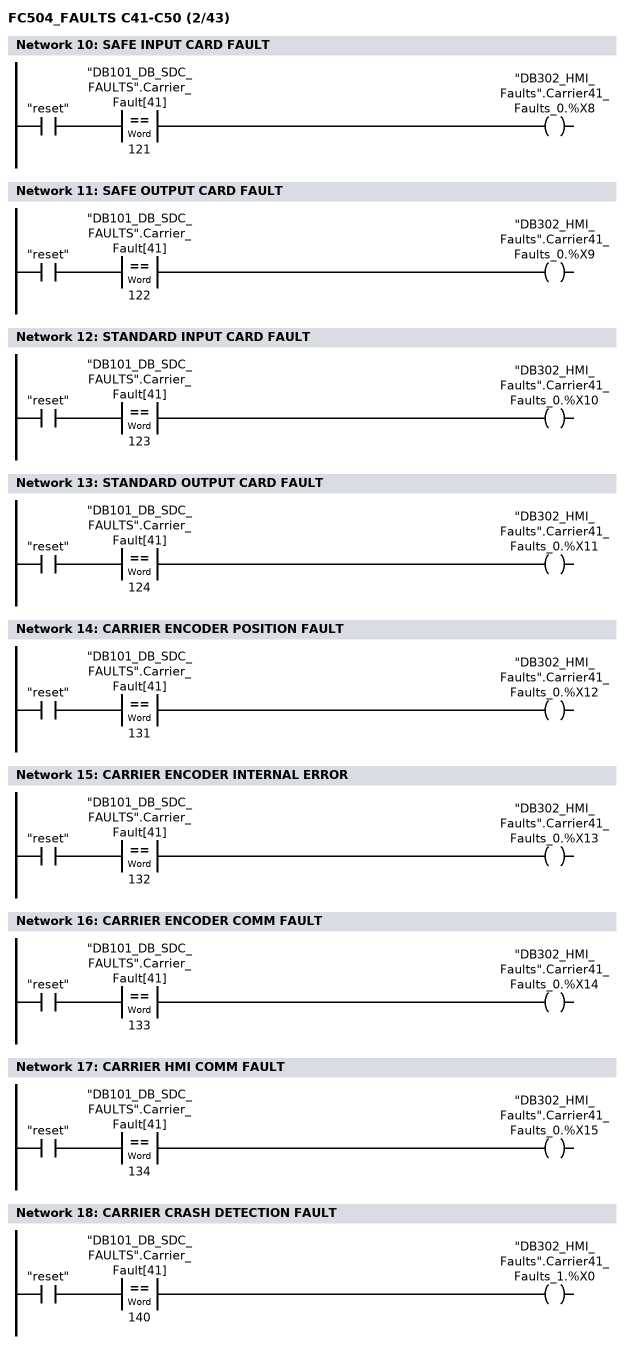
   RUNG wire#powerrail
      Contact( "reset" )
      { S7_Templates := "SrcType := Word" } EQ_Contact(in1 := "DB101_DB_SDC_FAULTS".Carrier_Fault[41], in2 := 121)
      Coil( "DB302_HMI_Faults".Carrier41_Faults_0.%X8 )
   END_RUNG
   // the same network as SCL:
   "DB302_HMI_Faults".Carrier41_Faults_0.%X8 := "reset" AND ("DB101_DB_SDC_FAULTS".Carrier_Fault[41] = 121);
END_REGION

REGION Network 11: SAFE OUTPUT CARD FAULT
   RUNG wire#powerrail
      Contact( "reset" )
      { S7_Templates := "SrcType := Word" } EQ_Contact(in1 := "DB101_DB_SDC_FAULTS".Carrier_Fault[41], in2 := 122)
      Coil( "DB302_HMI_Faults".Carrier41_Faults_0.%X9 )
   END_RUNG
   // the same network as SCL:
   "DB302_HMI_Faults".Carrier41_Faults_0.%X9 := "reset" AND ("DB101_DB_SDC_FAULTS".Carrier_Fault[41] = 122);
END_REGION

REGION Network 12: STANDARD INPUT CARD FAULT
   RUNG wire#powerrail
      Contact( "reset" )
      { S7_Templates := "SrcType := Word" } EQ_Contact(in1 := "DB101_DB_SDC_FAULTS".Carrier_Fault[41], in2 := 123)
      Coil( "DB302_HMI_Faults".Carrier41_Faults_0.%X10 )
   END_RUNG
   // the same network as SCL:
   "DB302_HMI_Faults".Carrier41_Faults_0.%X10 := "reset" AND ("DB101_DB_SDC_FAULTS".Carrier_Fault[41] = 123);
END_REGION

REGION Network 13: STANDARD OUTPUT CARD FAULT
   RUNG wire#powerrail
      Contact( "reset" )
      { S7_Templates := "SrcType := Word" } EQ_Contact(in1 := "DB101_DB_SDC_FAULTS".Carrier_Fault[41], in2 := 124)
      Coil( "DB302_HMI_Faults".Carrier41_Faults_0.%X11 )
   END_RUNG
   // the same network as SCL:
   "DB302_HMI_Faults".Carrier41_Faults_0.%X11 := "reset" AND ("DB101_DB_SDC_FAULTS".Carrier_Fault[41] = 124);
END_REGION

REGION Network 14: CARRIER ENCODER POSITION FAULT
   RUNG wire#powerrail
      Contact( "reset" )
      { S7_Templates := "SrcType := Word" } EQ_Contact(in1 := "DB101_DB_SDC_FAULTS".Carrier_Fault[41], in2 := 131)
      Coil( "DB302_HMI_Faults".Carrier41_Faults_0.%X12 )
   END_RUNG
   // the same network as SCL:
   "DB302_HMI_Faults".Carrier41_Faults_0.%X12 := "reset" AND ("DB101_DB_SDC_FAULTS".Carrier_Fault[41] = 131);
END_REGION

REGION Network 15: CARRIER ENCODER INTERNAL ERROR
   RUNG wire#powerrail
      Contact( "reset" )
      { S7_Templates := "SrcType := Word" } EQ_Contact(in1 := "DB101_DB_SDC_FAULTS".Carrier_Fault[41], in2 := 132)
      Coil( "DB302_HMI_Faults".Carrier41_Faults_0.%X13 )
   END_RUNG
   // the same network as SCL:
   "DB302_HMI_Faults".Carrier41_Faults_0.%X13 := "reset" AND ("DB101_DB_SDC_FAULTS".Carrier_Fault[41] = 132);
END_REGION

REGION Network 16: CARRIER ENCODER COMM FAULT
   RUNG wire#powerrail
      Contact( "reset" )
      { S7_Templates := "SrcType := Word" } EQ_Contact(in1 := "DB101_DB_SDC_FAULTS".Carrier_Fault[41], in2 := 133)
      Coil( "DB302_HMI_Faults".Carrier41_Faults_0.%X14 )
   END_RUNG
   // the same network as SCL:
   "DB302_HMI_Faults".Carrier41_Faults_0.%X14 := "reset" AND ("DB101_DB_SDC_FAULTS".Carrier_Fault[41] = 133);
END_REGION

REGION Network 17: CARRIER HMI COMM FAULT
   RUNG wire#powerrail
      Contact( "reset" )
      { S7_Templates := "SrcType := Word" } EQ_Contact(in1 := "DB101_DB_SDC_FAULTS".Carrier_Fault[41], in2 := 134)
      Coil( "DB302_HMI_Faults".Carrier41_Faults_0.%X15 )
   END_RUNG
   // the same network as SCL:
   "DB302_HMI_Faults".Carrier41_Faults_0.%X15 := "reset" AND ("DB101_DB_SDC_FAULTS".Carrier_Fault[41] = 134);
END_REGION

REGION Network 18: CARRIER CRASH DETECTION FAULT
   RUNG wire#powerrail
      Contact( "reset" )
      { S7_Templates := "SrcType := Word" } EQ_Contact(in1 := "DB101_DB_SDC_FAULTS".Carrier_Fault[41], in2 := 140)
      Coil( "DB302_HMI_Faults".Carrier41_Faults_1.%X0 )
   END_RUNG
   // the same network as SCL:
   "DB302_HMI_Faults".Carrier41_Faults_1.%X0 := "reset" AND ("DB101_DB_SDC_FAULTS".Carrier_Fault[41] = 140);
END_REGION

REGION Network 19: CARRIER NUMBER INVALID FAULT
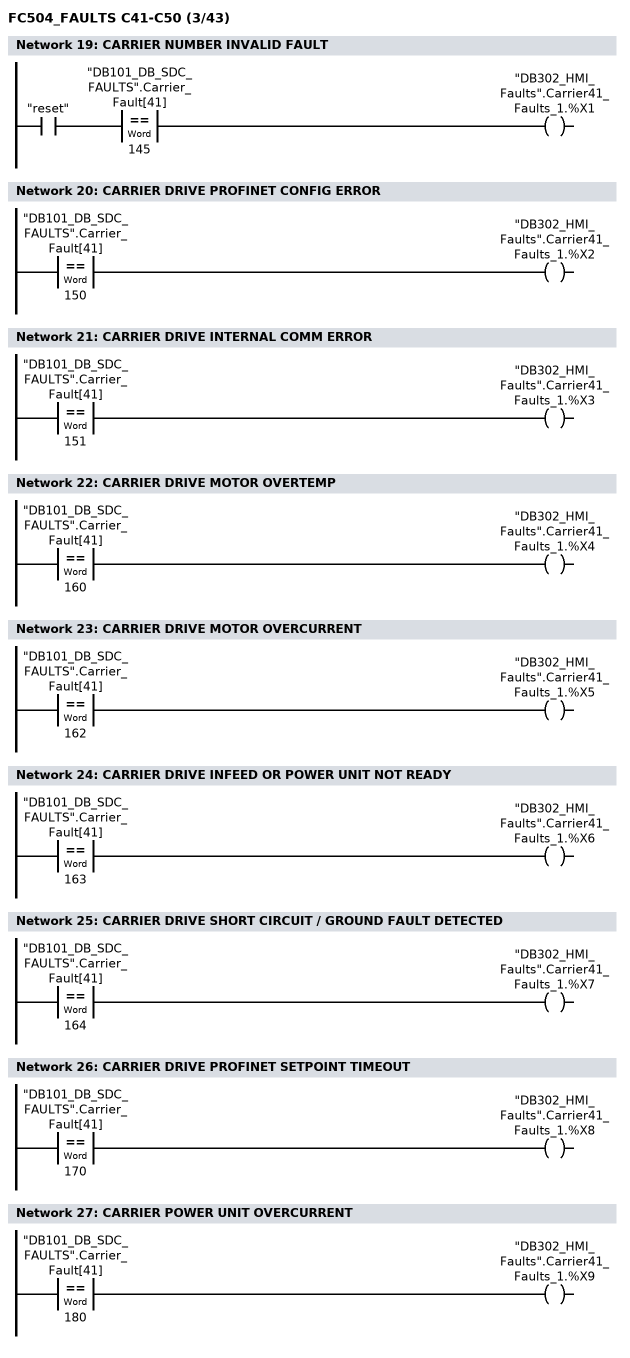
   RUNG wire#powerrail
      Contact( "reset" )
      { S7_Templates := "SrcType := Word" } EQ_Contact(in1 := "DB101_DB_SDC_FAULTS".Carrier_Fault[41], in2 := 145)
      Coil( "DB302_HMI_Faults".Carrier41_Faults_1.%X1 )
   END_RUNG
   // the same network as SCL:
   "DB302_HMI_Faults".Carrier41_Faults_1.%X1 := "reset" AND ("DB101_DB_SDC_FAULTS".Carrier_Fault[41] = 145);
END_REGION

REGION Network 20: CARRIER DRIVE PROFINET CONFIG ERROR
   RUNG wire#powerrail
      { S7_Templates := "SrcType := Word" } EQ_Contact(in1 := "DB101_DB_SDC_FAULTS".Carrier_Fault[41], in2 := 150)
      Coil( "DB302_HMI_Faults".Carrier41_Faults_1.%X2 )
   END_RUNG
   // the same network as SCL:
   "DB302_HMI_Faults".Carrier41_Faults_1.%X2 := "DB101_DB_SDC_FAULTS".Carrier_Fault[41] = 150;
END_REGION

REGION Network 21: CARRIER DRIVE INTERNAL COMM ERROR
   RUNG wire#powerrail
      { S7_Templates := "SrcType := Word" } EQ_Contact(in1 := "DB101_DB_SDC_FAULTS".Carrier_Fault[41], in2 := 151)
      Coil( "DB302_HMI_Faults".Carrier41_Faults_1.%X3 )
   END_RUNG
   // the same network as SCL:
   "DB302_HMI_Faults".Carrier41_Faults_1.%X3 := "DB101_DB_SDC_FAULTS".Carrier_Fault[41] = 151;
END_REGION

REGION Network 22: CARRIER DRIVE MOTOR OVERTEMP
   RUNG wire#powerrail
      { S7_Templates := "SrcType := Word" } EQ_Contact(in1 := "DB101_DB_SDC_FAULTS".Carrier_Fault[41], in2 := 160)
      Coil( "DB302_HMI_Faults".Carrier41_Faults_1.%X4 )
   END_RUNG
   // the same network as SCL:
   "DB302_HMI_Faults".Carrier41_Faults_1.%X4 := "DB101_DB_SDC_FAULTS".Carrier_Fault[41] = 160;
END_REGION

REGION Network 23: CARRIER DRIVE MOTOR OVERCURRENT
   RUNG wire#powerrail
      { S7_Templates := "SrcType := Word" } EQ_Contact(in1 := "DB101_DB_SDC_FAULTS".Carrier_Fault[41], in2 := 162)
      Coil( "DB302_HMI_Faults".Carrier41_Faults_1.%X5 )
   END_RUNG
   // the same network as SCL:
   "DB302_HMI_Faults".Carrier41_Faults_1.%X5 := "DB101_DB_SDC_FAULTS".Carrier_Fault[41] = 162;
END_REGION

REGION Network 24: CARRIER DRIVE INFEED OR POWER UNIT NOT READY
   RUNG wire#powerrail
      { S7_Templates := "SrcType := Word" } EQ_Contact(in1 := "DB101_DB_SDC_FAULTS".Carrier_Fault[41], in2 := 163)
      Coil( "DB302_HMI_Faults".Carrier41_Faults_1.%X6 )
   END_RUNG
   // the same network as SCL:
   "DB302_HMI_Faults".Carrier41_Faults_1.%X6 := "DB101_DB_SDC_FAULTS".Carrier_Fault[41] = 163;
END_REGION

REGION Network 25: CARRIER DRIVE SHORT CIRCUIT / GROUND FAULT DETECTED
   RUNG wire#powerrail
      { S7_Templates := "SrcType := Word" } EQ_Contact(in1 := "DB101_DB_SDC_FAULTS".Carrier_Fault[41], in2 := 164)
      Coil( "DB302_HMI_Faults".Carrier41_Faults_1.%X7 )
   END_RUNG
   // the same network as SCL:
   "DB302_HMI_Faults".Carrier41_Faults_1.%X7 := "DB101_DB_SDC_FAULTS".Carrier_Fault[41] = 164;
END_REGION

REGION Network 26: CARRIER DRIVE PROFINET SETPOINT TIMEOUT
   RUNG wire#powerrail
      { S7_Templates := "SrcType := Word" } EQ_Contact(in1 := "DB101_DB_SDC_FAULTS".Carrier_Fault[41], in2 := 170)
      Coil( "DB302_HMI_Faults".Carrier41_Faults_1.%X8 )
   END_RUNG
   // the same network as SCL:
   "DB302_HMI_Faults".Carrier41_Faults_1.%X8 := "DB101_DB_SDC_FAULTS".Carrier_Fault[41] = 170;
END_REGION

REGION Network 27: CARRIER POWER UNIT OVERCURRENT
   RUNG wire#powerrail
      { S7_Templates := "SrcType := Word" } EQ_Contact(in1 := "DB101_DB_SDC_FAULTS".Carrier_Fault[41], in2 := 180)
      Coil( "DB302_HMI_Faults".Carrier41_Faults_1.%X9 )
   END_RUNG
   // the same network as SCL:
   "DB302_HMI_Faults".Carrier41_Faults_1.%X9 := "DB101_DB_SDC_FAULTS".Carrier_Fault[41] = 180;
END_REGION

REGION Network 28: CARRIER POWER UNIT DC LINK OVERVOLTAGE
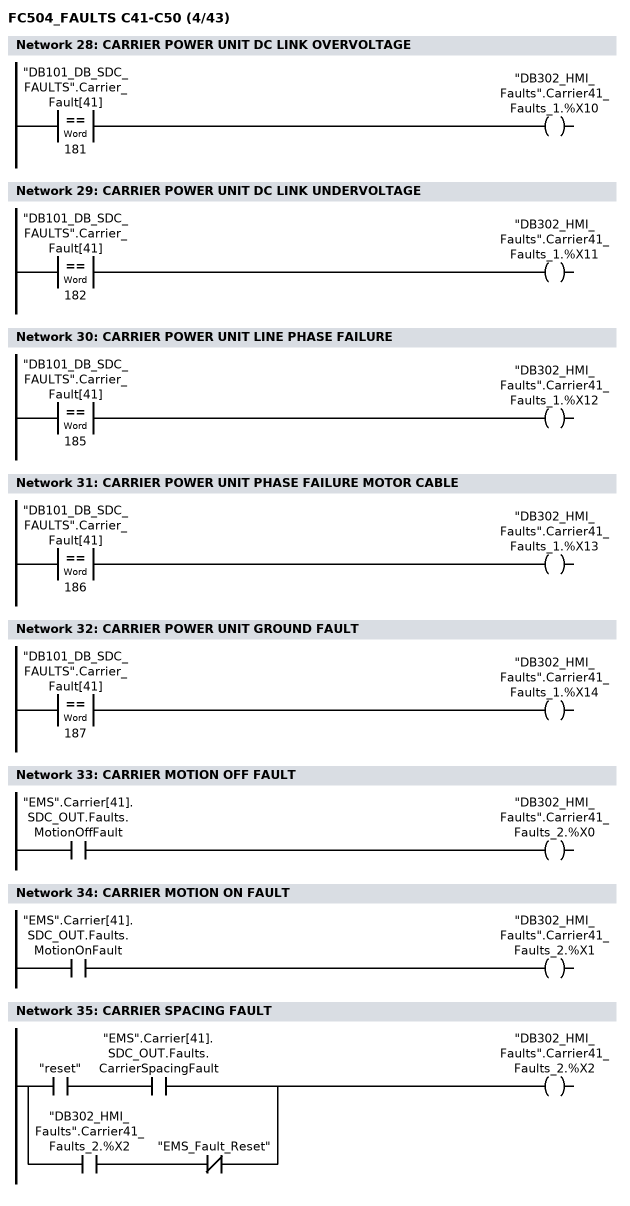
   RUNG wire#powerrail
      { S7_Templates := "SrcType := Word" } EQ_Contact(in1 := "DB101_DB_SDC_FAULTS".Carrier_Fault[41], in2 := 181)
      Coil( "DB302_HMI_Faults".Carrier41_Faults_1.%X10 )
   END_RUNG
   // the same network as SCL:
   "DB302_HMI_Faults".Carrier41_Faults_1.%X10 := "DB101_DB_SDC_FAULTS".Carrier_Fault[41] = 181;
END_REGION

REGION Network 29: CARRIER POWER UNIT DC LINK UNDERVOLTAGE
   RUNG wire#powerrail
      { S7_Templates := "SrcType := Word" } EQ_Contact(in1 := "DB101_DB_SDC_FAULTS".Carrier_Fault[41], in2 := 182)
      Coil( "DB302_HMI_Faults".Carrier41_Faults_1.%X11 )
   END_RUNG
   // the same network as SCL:
   "DB302_HMI_Faults".Carrier41_Faults_1.%X11 := "DB101_DB_SDC_FAULTS".Carrier_Fault[41] = 182;
END_REGION

REGION Network 30: CARRIER POWER UNIT LINE PHASE FAILURE
   RUNG wire#powerrail
      { S7_Templates := "SrcType := Word" } EQ_Contact(in1 := "DB101_DB_SDC_FAULTS".Carrier_Fault[41], in2 := 185)
      Coil( "DB302_HMI_Faults".Carrier41_Faults_1.%X12 )
   END_RUNG
   // the same network as SCL:
   "DB302_HMI_Faults".Carrier41_Faults_1.%X12 := "DB101_DB_SDC_FAULTS".Carrier_Fault[41] = 185;
END_REGION

REGION Network 31: CARRIER POWER UNIT PHASE FAILURE MOTOR CABLE
   RUNG wire#powerrail
      { S7_Templates := "SrcType := Word" } EQ_Contact(in1 := "DB101_DB_SDC_FAULTS".Carrier_Fault[41], in2 := 186)
      Coil( "DB302_HMI_Faults".Carrier41_Faults_1.%X13 )
   END_RUNG
   // the same network as SCL:
   "DB302_HMI_Faults".Carrier41_Faults_1.%X13 := "DB101_DB_SDC_FAULTS".Carrier_Fault[41] = 186;
END_REGION

REGION Network 32: CARRIER POWER UNIT GROUND FAULT
   RUNG wire#powerrail
      { S7_Templates := "SrcType := Word" } EQ_Contact(in1 := "DB101_DB_SDC_FAULTS".Carrier_Fault[41], in2 := 187)
      Coil( "DB302_HMI_Faults".Carrier41_Faults_1.%X14 )
   END_RUNG
   // the same network as SCL:
   "DB302_HMI_Faults".Carrier41_Faults_1.%X14 := "DB101_DB_SDC_FAULTS".Carrier_Fault[41] = 187;
END_REGION

REGION Network 33: CARRIER MOTION OFF FAULT
   RUNG wire#powerrail
      Contact( "EMS".Carrier[41].SDC_OUT.Faults.MotionOffFault )
      Coil( "DB302_HMI_Faults".Carrier41_Faults_2.%X0 )
   END_RUNG
   // the same network as SCL:
   "DB302_HMI_Faults".Carrier41_Faults_2.%X0 := "EMS".Carrier[41].SDC_OUT.Faults.MotionOffFault;
END_REGION

REGION Network 34: CARRIER MOTION ON FAULT
   RUNG wire#powerrail
      Contact( "EMS".Carrier[41].SDC_OUT.Faults.MotionOnFault )
      Coil( "DB302_HMI_Faults".Carrier41_Faults_2.%X1 )
   END_RUNG
   // the same network as SCL:
   "DB302_HMI_Faults".Carrier41_Faults_2.%X1 := "EMS".Carrier[41].SDC_OUT.Faults.MotionOnFault;
END_REGION

REGION Network 35: CARRIER SPACING FAULT
   RUNG wire#powerrail
      Contact( "reset" )
      Contact( "EMS".Carrier[41].SDC_OUT.Faults.CarrierSpacingFault )
      wire#w1
      Coil( "DB302_HMI_Faults".Carrier41_Faults_2.%X2 )
   END_RUNG
   RUNG wire#powerrail
      Contact( "DB302_HMI_Faults".Carrier41_Faults_2.%X2 )
      I_Contact( "EMS_Fault_Reset" )
   END_RUNG wire#w1
   // the same network as SCL:
   "DB302_HMI_Faults".Carrier41_Faults_2.%X2 := ("reset" AND "EMS".Carrier[41].SDC_OUT.Faults.CarrierSpacingFault) OR ("DB302_HMI_Faults".Carrier41_Faults_2.%X2 AND NOT "EMS_Fault_Reset");
END_REGION

REGION Network 36: DUPLICATE CARRIER NUMBER FAULT
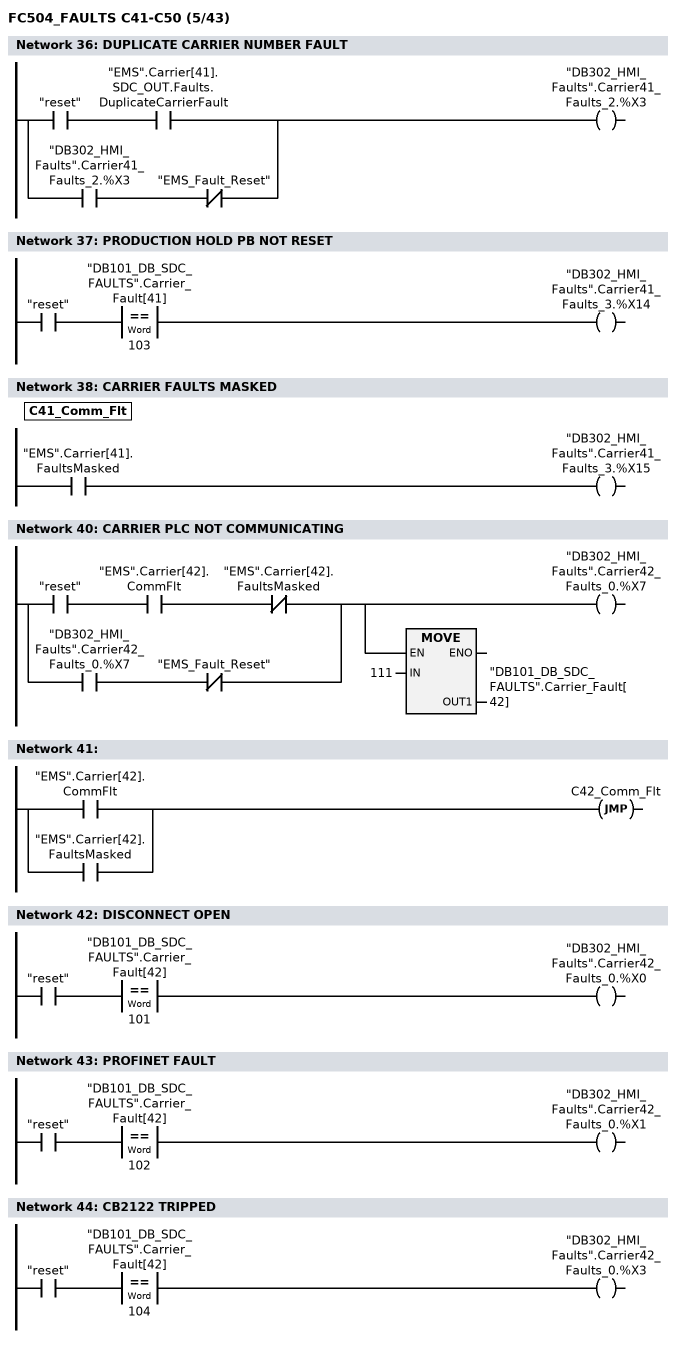
   RUNG wire#powerrail
      Contact( "reset" )
      Contact( "EMS".Carrier[41].SDC_OUT.Faults.DuplicateCarrierFault )
      wire#w1
      Coil( "DB302_HMI_Faults".Carrier41_Faults_2.%X3 )
   END_RUNG
   RUNG wire#powerrail
      Contact( "DB302_HMI_Faults".Carrier41_Faults_2.%X3 )
      I_Contact( "EMS_Fault_Reset" )
   END_RUNG wire#w1
   // the same network as SCL:
   "DB302_HMI_Faults".Carrier41_Faults_2.%X3 := ("reset" AND "EMS".Carrier[41].SDC_OUT.Faults.DuplicateCarrierFault) OR ("DB302_HMI_Faults".Carrier41_Faults_2.%X3 AND NOT "EMS_Fault_Reset");
END_REGION

REGION Network 37: PRODUCTION HOLD PB NOT RESET
   RUNG wire#powerrail
      Contact( "reset" )
      { S7_Templates := "SrcType := Word" } EQ_Contact(in1 := "DB101_DB_SDC_FAULTS".Carrier_Fault[41], in2 := 103)
      Coil( "DB302_HMI_Faults".Carrier41_Faults_3.%X14 )
   END_RUNG
   // the same network as SCL:
   "DB302_HMI_Faults".Carrier41_Faults_3.%X14 := "reset" AND ("DB101_DB_SDC_FAULTS".Carrier_Fault[41] = 103);
END_REGION

REGION Network 38: CARRIER FAULTS MASKED
   Label( C41_Comm_Flt )
   RUNG wire#powerrail
      Contact( "EMS".Carrier[41].FaultsMasked )
      Coil( "DB302_HMI_Faults".Carrier41_Faults_3.%X15 )
   END_RUNG
   // the same network as SCL:
   C41_Comm_Flt:
   "DB302_HMI_Faults".Carrier41_Faults_3.%X15 := "EMS".Carrier[41].FaultsMasked;
END_REGION

REGION Network 39: CARRIER 42 FAULTS
END_REGION

REGION Network 40: CARRIER PLC NOT COMMUNICATING
   RUNG wire#powerrail
      Contact( "reset" )
      Contact( "EMS".Carrier[42].CommFlt )
      I_Contact( "EMS".Carrier[42].FaultsMasked )
      wire#w1
      Coil( "DB302_HMI_Faults".Carrier42_Faults_0.%X7 )
   END_RUNG
   RUNG wire#powerrail
      Contact( "DB302_HMI_Faults".Carrier42_Faults_0.%X7 )
      I_Contact( "EMS_Fault_Reset" )
   END_RUNG wire#w1
   RUNG wire#w1
      Move(in := 111, out1 => "DB101_DB_SDC_FAULTS".Carrier_Fault[42])
   END_RUNG
   // the same network as SCL:
   "DB302_HMI_Faults".Carrier42_Faults_0.%X7 := ("reset" AND "EMS".Carrier[42].CommFlt AND NOT "EMS".Carrier[42].FaultsMasked) OR ("DB302_HMI_Faults".Carrier42_Faults_0.%X7 AND NOT "EMS_Fault_Reset");
   IF "DB302_HMI_Faults".Carrier42_Faults_0.%X7 THEN "DB101_DB_SDC_FAULTS".Carrier_Fault[42] := 111; END_IF;
END_REGION

REGION Network 41
   RUNG wire#powerrail
      Contact( "EMS".Carrier[42].CommFlt )
      wire#w1
      JumpCoil( C42_Comm_Flt )
   END_RUNG
   RUNG wire#powerrail
      Contact( "EMS".Carrier[42].FaultsMasked )
   END_RUNG wire#w1
   // the same network as SCL:
   IF "EMS".Carrier[42].CommFlt OR "EMS".Carrier[42].FaultsMasked THEN GOTO C42_Comm_Flt; END_IF;
END_REGION

REGION Network 42: DISCONNECT OPEN
   RUNG wire#powerrail
      Contact( "reset" )
      { S7_Templates := "SrcType := Word" } EQ_Contact(in1 := "DB101_DB_SDC_FAULTS".Carrier_Fault[42], in2 := 101)
      Coil( "DB302_HMI_Faults".Carrier42_Faults_0.%X0 )
   END_RUNG
   // the same network as SCL:
   "DB302_HMI_Faults".Carrier42_Faults_0.%X0 := "reset" AND ("DB101_DB_SDC_FAULTS".Carrier_Fault[42] = 101);
END_REGION

REGION Network 43: PROFINET FAULT
   RUNG wire#powerrail
      Contact( "reset" )
      { S7_Templates := "SrcType := Word" } EQ_Contact(in1 := "DB101_DB_SDC_FAULTS".Carrier_Fault[42], in2 := 102)
      Coil( "DB302_HMI_Faults".Carrier42_Faults_0.%X1 )
   END_RUNG
   // the same network as SCL:
   "DB302_HMI_Faults".Carrier42_Faults_0.%X1 := "reset" AND ("DB101_DB_SDC_FAULTS".Carrier_Fault[42] = 102);
END_REGION

REGION Network 44: CB2122 TRIPPED
   RUNG wire#powerrail
      Contact( "reset" )
      { S7_Templates := "SrcType := Word" } EQ_Contact(in1 := "DB101_DB_SDC_FAULTS".Carrier_Fault[42], in2 := 104)
      Coil( "DB302_HMI_Faults".Carrier42_Faults_0.%X3 )
   END_RUNG
   // the same network as SCL:
   "DB302_HMI_Faults".Carrier42_Faults_0.%X3 := "reset" AND ("DB101_DB_SDC_FAULTS".Carrier_Fault[42] = 104);
END_REGION

REGION Network 45: CB2123 TRIPPED
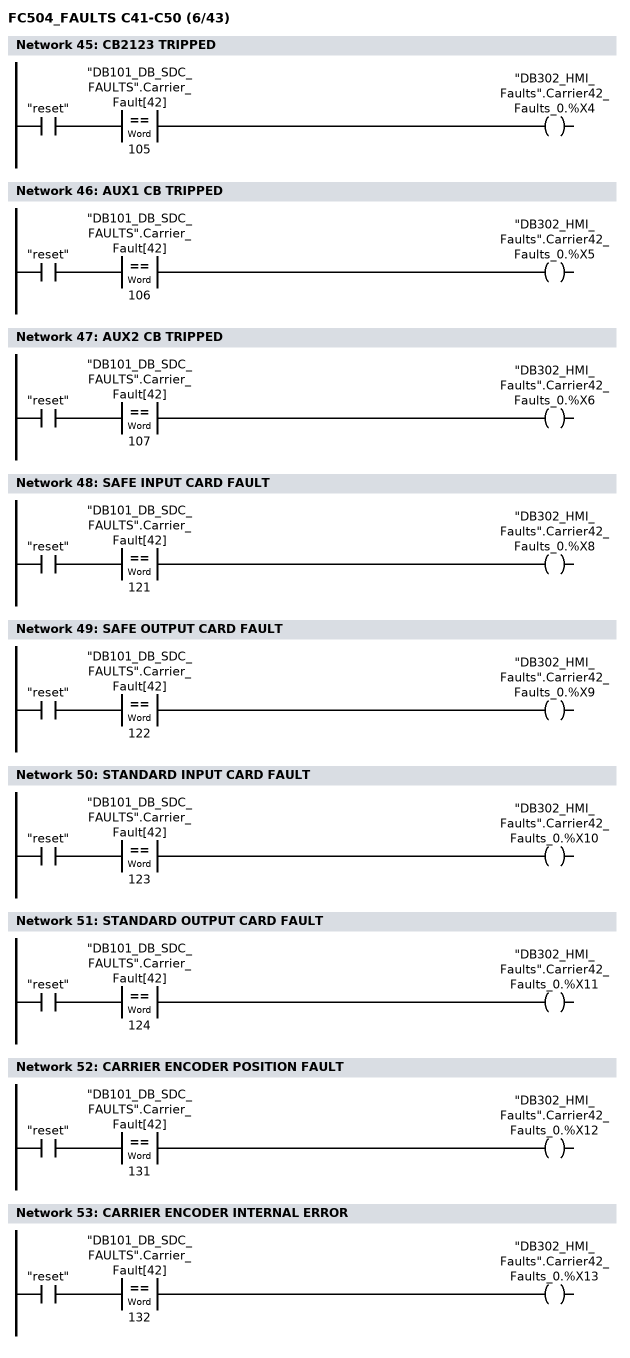
   RUNG wire#powerrail
      Contact( "reset" )
      { S7_Templates := "SrcType := Word" } EQ_Contact(in1 := "DB101_DB_SDC_FAULTS".Carrier_Fault[42], in2 := 105)
      Coil( "DB302_HMI_Faults".Carrier42_Faults_0.%X4 )
   END_RUNG
   // the same network as SCL:
   "DB302_HMI_Faults".Carrier42_Faults_0.%X4 := "reset" AND ("DB101_DB_SDC_FAULTS".Carrier_Fault[42] = 105);
END_REGION

REGION Network 46: AUX1 CB TRIPPED
   RUNG wire#powerrail
      Contact( "reset" )
      { S7_Templates := "SrcType := Word" } EQ_Contact(in1 := "DB101_DB_SDC_FAULTS".Carrier_Fault[42], in2 := 106)
      Coil( "DB302_HMI_Faults".Carrier42_Faults_0.%X5 )
   END_RUNG
   // the same network as SCL:
   "DB302_HMI_Faults".Carrier42_Faults_0.%X5 := "reset" AND ("DB101_DB_SDC_FAULTS".Carrier_Fault[42] = 106);
END_REGION

REGION Network 47: AUX2 CB TRIPPED
   RUNG wire#powerrail
      Contact( "reset" )
      { S7_Templates := "SrcType := Word" } EQ_Contact(in1 := "DB101_DB_SDC_FAULTS".Carrier_Fault[42], in2 := 107)
      Coil( "DB302_HMI_Faults".Carrier42_Faults_0.%X6 )
   END_RUNG
   // the same network as SCL:
   "DB302_HMI_Faults".Carrier42_Faults_0.%X6 := "reset" AND ("DB101_DB_SDC_FAULTS".Carrier_Fault[42] = 107);
END_REGION

REGION Network 48: SAFE INPUT CARD FAULT
   RUNG wire#powerrail
      Contact( "reset" )
      { S7_Templates := "SrcType := Word" } EQ_Contact(in1 := "DB101_DB_SDC_FAULTS".Carrier_Fault[42], in2 := 121)
      Coil( "DB302_HMI_Faults".Carrier42_Faults_0.%X8 )
   END_RUNG
   // the same network as SCL:
   "DB302_HMI_Faults".Carrier42_Faults_0.%X8 := "reset" AND ("DB101_DB_SDC_FAULTS".Carrier_Fault[42] = 121);
END_REGION

REGION Network 49: SAFE OUTPUT CARD FAULT
   RUNG wire#powerrail
      Contact( "reset" )
      { S7_Templates := "SrcType := Word" } EQ_Contact(in1 := "DB101_DB_SDC_FAULTS".Carrier_Fault[42], in2 := 122)
      Coil( "DB302_HMI_Faults".Carrier42_Faults_0.%X9 )
   END_RUNG
   // the same network as SCL:
   "DB302_HMI_Faults".Carrier42_Faults_0.%X9 := "reset" AND ("DB101_DB_SDC_FAULTS".Carrier_Fault[42] = 122);
END_REGION

REGION Network 50: STANDARD INPUT CARD FAULT
   RUNG wire#powerrail
      Contact( "reset" )
      { S7_Templates := "SrcType := Word" } EQ_Contact(in1 := "DB101_DB_SDC_FAULTS".Carrier_Fault[42], in2 := 123)
      Coil( "DB302_HMI_Faults".Carrier42_Faults_0.%X10 )
   END_RUNG
   // the same network as SCL:
   "DB302_HMI_Faults".Carrier42_Faults_0.%X10 := "reset" AND ("DB101_DB_SDC_FAULTS".Carrier_Fault[42] = 123);
END_REGION

REGION Network 51: STANDARD OUTPUT CARD FAULT
   RUNG wire#powerrail
      Contact( "reset" )
      { S7_Templates := "SrcType := Word" } EQ_Contact(in1 := "DB101_DB_SDC_FAULTS".Carrier_Fault[42], in2 := 124)
      Coil( "DB302_HMI_Faults".Carrier42_Faults_0.%X11 )
   END_RUNG
   // the same network as SCL:
   "DB302_HMI_Faults".Carrier42_Faults_0.%X11 := "reset" AND ("DB101_DB_SDC_FAULTS".Carrier_Fault[42] = 124);
END_REGION

REGION Network 52: CARRIER ENCODER POSITION FAULT
   RUNG wire#powerrail
      Contact( "reset" )
      { S7_Templates := "SrcType := Word" } EQ_Contact(in1 := "DB101_DB_SDC_FAULTS".Carrier_Fault[42], in2 := 131)
      Coil( "DB302_HMI_Faults".Carrier42_Faults_0.%X12 )
   END_RUNG
   // the same network as SCL:
   "DB302_HMI_Faults".Carrier42_Faults_0.%X12 := "reset" AND ("DB101_DB_SDC_FAULTS".Carrier_Fault[42] = 131);
END_REGION

REGION Network 53: CARRIER ENCODER INTERNAL ERROR
   RUNG wire#powerrail
      Contact( "reset" )
      { S7_Templates := "SrcType := Word" } EQ_Contact(in1 := "DB101_DB_SDC_FAULTS".Carrier_Fault[42], in2 := 132)
      Coil( "DB302_HMI_Faults".Carrier42_Faults_0.%X13 )
   END_RUNG
   // the same network as SCL:
   "DB302_HMI_Faults".Carrier42_Faults_0.%X13 := "reset" AND ("DB101_DB_SDC_FAULTS".Carrier_Fault[42] = 132);
END_REGION

REGION Network 54: CARRIER ENCODER COMM FAULT
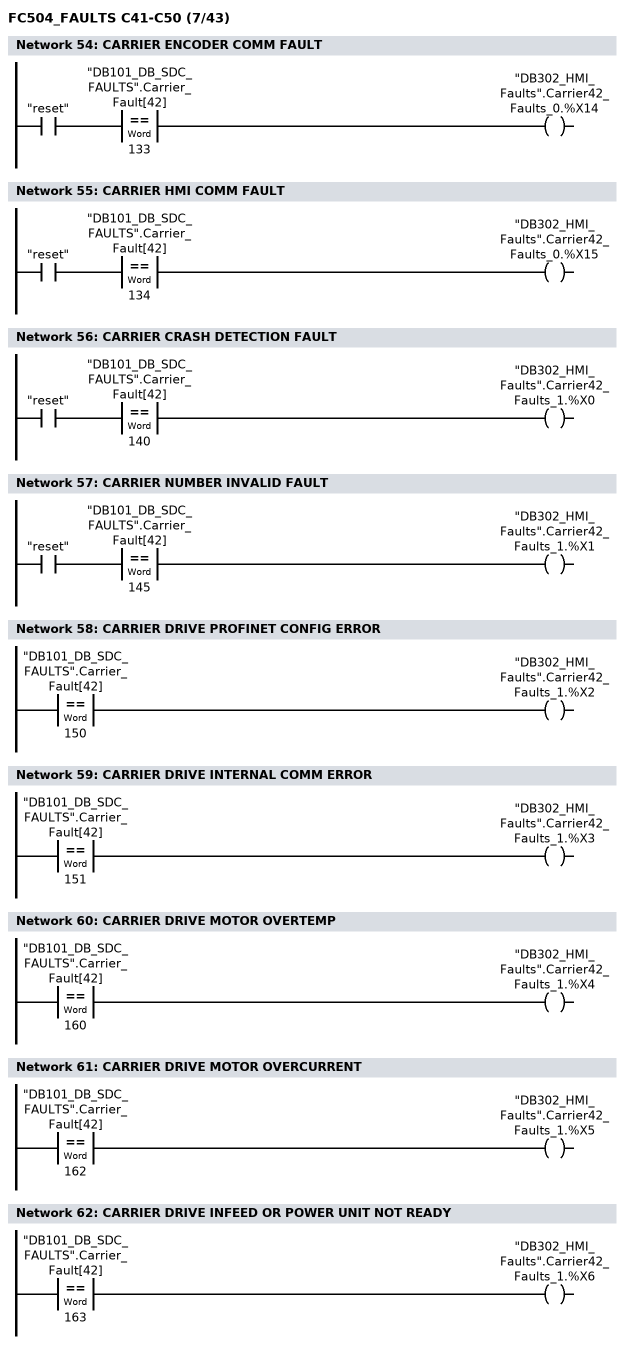
   RUNG wire#powerrail
      Contact( "reset" )
      { S7_Templates := "SrcType := Word" } EQ_Contact(in1 := "DB101_DB_SDC_FAULTS".Carrier_Fault[42], in2 := 133)
      Coil( "DB302_HMI_Faults".Carrier42_Faults_0.%X14 )
   END_RUNG
   // the same network as SCL:
   "DB302_HMI_Faults".Carrier42_Faults_0.%X14 := "reset" AND ("DB101_DB_SDC_FAULTS".Carrier_Fault[42] = 133);
END_REGION

REGION Network 55: CARRIER HMI COMM FAULT
   RUNG wire#powerrail
      Contact( "reset" )
      { S7_Templates := "SrcType := Word" } EQ_Contact(in1 := "DB101_DB_SDC_FAULTS".Carrier_Fault[42], in2 := 134)
      Coil( "DB302_HMI_Faults".Carrier42_Faults_0.%X15 )
   END_RUNG
   // the same network as SCL:
   "DB302_HMI_Faults".Carrier42_Faults_0.%X15 := "reset" AND ("DB101_DB_SDC_FAULTS".Carrier_Fault[42] = 134);
END_REGION

REGION Network 56: CARRIER CRASH DETECTION FAULT
   RUNG wire#powerrail
      Contact( "reset" )
      { S7_Templates := "SrcType := Word" } EQ_Contact(in1 := "DB101_DB_SDC_FAULTS".Carrier_Fault[42], in2 := 140)
      Coil( "DB302_HMI_Faults".Carrier42_Faults_1.%X0 )
   END_RUNG
   // the same network as SCL:
   "DB302_HMI_Faults".Carrier42_Faults_1.%X0 := "reset" AND ("DB101_DB_SDC_FAULTS".Carrier_Fault[42] = 140);
END_REGION

REGION Network 57: CARRIER NUMBER INVALID FAULT
   RUNG wire#powerrail
      Contact( "reset" )
      { S7_Templates := "SrcType := Word" } EQ_Contact(in1 := "DB101_DB_SDC_FAULTS".Carrier_Fault[42], in2 := 145)
      Coil( "DB302_HMI_Faults".Carrier42_Faults_1.%X1 )
   END_RUNG
   // the same network as SCL:
   "DB302_HMI_Faults".Carrier42_Faults_1.%X1 := "reset" AND ("DB101_DB_SDC_FAULTS".Carrier_Fault[42] = 145);
END_REGION

REGION Network 58: CARRIER DRIVE PROFINET CONFIG ERROR
   RUNG wire#powerrail
      { S7_Templates := "SrcType := Word" } EQ_Contact(in1 := "DB101_DB_SDC_FAULTS".Carrier_Fault[42], in2 := 150)
      Coil( "DB302_HMI_Faults".Carrier42_Faults_1.%X2 )
   END_RUNG
   // the same network as SCL:
   "DB302_HMI_Faults".Carrier42_Faults_1.%X2 := "DB101_DB_SDC_FAULTS".Carrier_Fault[42] = 150;
END_REGION

REGION Network 59: CARRIER DRIVE INTERNAL COMM ERROR
   RUNG wire#powerrail
      { S7_Templates := "SrcType := Word" } EQ_Contact(in1 := "DB101_DB_SDC_FAULTS".Carrier_Fault[42], in2 := 151)
      Coil( "DB302_HMI_Faults".Carrier42_Faults_1.%X3 )
   END_RUNG
   // the same network as SCL:
   "DB302_HMI_Faults".Carrier42_Faults_1.%X3 := "DB101_DB_SDC_FAULTS".Carrier_Fault[42] = 151;
END_REGION

REGION Network 60: CARRIER DRIVE MOTOR OVERTEMP
   RUNG wire#powerrail
      { S7_Templates := "SrcType := Word" } EQ_Contact(in1 := "DB101_DB_SDC_FAULTS".Carrier_Fault[42], in2 := 160)
      Coil( "DB302_HMI_Faults".Carrier42_Faults_1.%X4 )
   END_RUNG
   // the same network as SCL:
   "DB302_HMI_Faults".Carrier42_Faults_1.%X4 := "DB101_DB_SDC_FAULTS".Carrier_Fault[42] = 160;
END_REGION

REGION Network 61: CARRIER DRIVE MOTOR OVERCURRENT
   RUNG wire#powerrail
      { S7_Templates := "SrcType := Word" } EQ_Contact(in1 := "DB101_DB_SDC_FAULTS".Carrier_Fault[42], in2 := 162)
      Coil( "DB302_HMI_Faults".Carrier42_Faults_1.%X5 )
   END_RUNG
   // the same network as SCL:
   "DB302_HMI_Faults".Carrier42_Faults_1.%X5 := "DB101_DB_SDC_FAULTS".Carrier_Fault[42] = 162;
END_REGION

REGION Network 62: CARRIER DRIVE INFEED OR POWER UNIT NOT READY
   RUNG wire#powerrail
      { S7_Templates := "SrcType := Word" } EQ_Contact(in1 := "DB101_DB_SDC_FAULTS".Carrier_Fault[42], in2 := 163)
      Coil( "DB302_HMI_Faults".Carrier42_Faults_1.%X6 )
   END_RUNG
   // the same network as SCL:
   "DB302_HMI_Faults".Carrier42_Faults_1.%X6 := "DB101_DB_SDC_FAULTS".Carrier_Fault[42] = 163;
END_REGION

REGION Network 63: CARRIER DRIVE SHORT CIRCUIT / GROUND FAULT DETECTED
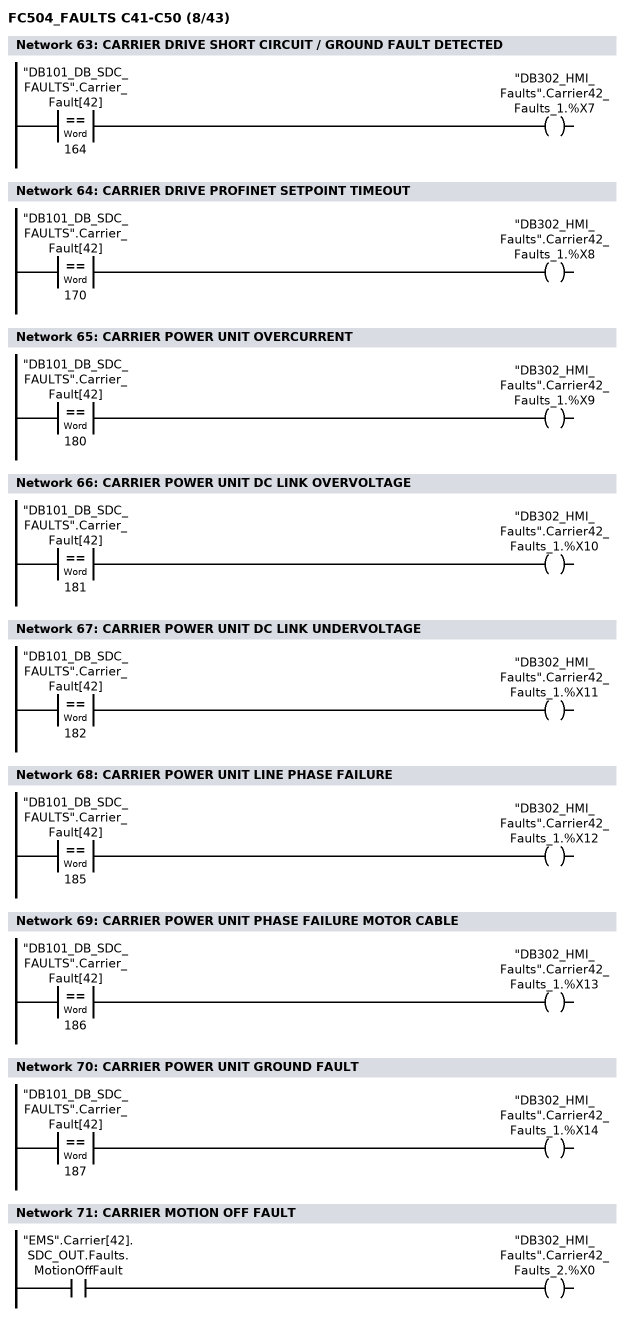
   RUNG wire#powerrail
      { S7_Templates := "SrcType := Word" } EQ_Contact(in1 := "DB101_DB_SDC_FAULTS".Carrier_Fault[42], in2 := 164)
      Coil( "DB302_HMI_Faults".Carrier42_Faults_1.%X7 )
   END_RUNG
   // the same network as SCL:
   "DB302_HMI_Faults".Carrier42_Faults_1.%X7 := "DB101_DB_SDC_FAULTS".Carrier_Fault[42] = 164;
END_REGION

REGION Network 64: CARRIER DRIVE PROFINET SETPOINT TIMEOUT
   RUNG wire#powerrail
      { S7_Templates := "SrcType := Word" } EQ_Contact(in1 := "DB101_DB_SDC_FAULTS".Carrier_Fault[42], in2 := 170)
      Coil( "DB302_HMI_Faults".Carrier42_Faults_1.%X8 )
   END_RUNG
   // the same network as SCL:
   "DB302_HMI_Faults".Carrier42_Faults_1.%X8 := "DB101_DB_SDC_FAULTS".Carrier_Fault[42] = 170;
END_REGION

REGION Network 65: CARRIER POWER UNIT OVERCURRENT
   RUNG wire#powerrail
      { S7_Templates := "SrcType := Word" } EQ_Contact(in1 := "DB101_DB_SDC_FAULTS".Carrier_Fault[42], in2 := 180)
      Coil( "DB302_HMI_Faults".Carrier42_Faults_1.%X9 )
   END_RUNG
   // the same network as SCL:
   "DB302_HMI_Faults".Carrier42_Faults_1.%X9 := "DB101_DB_SDC_FAULTS".Carrier_Fault[42] = 180;
END_REGION

REGION Network 66: CARRIER POWER UNIT DC LINK OVERVOLTAGE
   RUNG wire#powerrail
      { S7_Templates := "SrcType := Word" } EQ_Contact(in1 := "DB101_DB_SDC_FAULTS".Carrier_Fault[42], in2 := 181)
      Coil( "DB302_HMI_Faults".Carrier42_Faults_1.%X10 )
   END_RUNG
   // the same network as SCL:
   "DB302_HMI_Faults".Carrier42_Faults_1.%X10 := "DB101_DB_SDC_FAULTS".Carrier_Fault[42] = 181;
END_REGION

REGION Network 67: CARRIER POWER UNIT DC LINK UNDERVOLTAGE
   RUNG wire#powerrail
      { S7_Templates := "SrcType := Word" } EQ_Contact(in1 := "DB101_DB_SDC_FAULTS".Carrier_Fault[42], in2 := 182)
      Coil( "DB302_HMI_Faults".Carrier42_Faults_1.%X11 )
   END_RUNG
   // the same network as SCL:
   "DB302_HMI_Faults".Carrier42_Faults_1.%X11 := "DB101_DB_SDC_FAULTS".Carrier_Fault[42] = 182;
END_REGION

REGION Network 68: CARRIER POWER UNIT LINE PHASE FAILURE
   RUNG wire#powerrail
      { S7_Templates := "SrcType := Word" } EQ_Contact(in1 := "DB101_DB_SDC_FAULTS".Carrier_Fault[42], in2 := 185)
      Coil( "DB302_HMI_Faults".Carrier42_Faults_1.%X12 )
   END_RUNG
   // the same network as SCL:
   "DB302_HMI_Faults".Carrier42_Faults_1.%X12 := "DB101_DB_SDC_FAULTS".Carrier_Fault[42] = 185;
END_REGION

REGION Network 69: CARRIER POWER UNIT PHASE FAILURE MOTOR CABLE
   RUNG wire#powerrail
      { S7_Templates := "SrcType := Word" } EQ_Contact(in1 := "DB101_DB_SDC_FAULTS".Carrier_Fault[42], in2 := 186)
      Coil( "DB302_HMI_Faults".Carrier42_Faults_1.%X13 )
   END_RUNG
   // the same network as SCL:
   "DB302_HMI_Faults".Carrier42_Faults_1.%X13 := "DB101_DB_SDC_FAULTS".Carrier_Fault[42] = 186;
END_REGION

REGION Network 70: CARRIER POWER UNIT GROUND FAULT
   RUNG wire#powerrail
      { S7_Templates := "SrcType := Word" } EQ_Contact(in1 := "DB101_DB_SDC_FAULTS".Carrier_Fault[42], in2 := 187)
      Coil( "DB302_HMI_Faults".Carrier42_Faults_1.%X14 )
   END_RUNG
   // the same network as SCL:
   "DB302_HMI_Faults".Carrier42_Faults_1.%X14 := "DB101_DB_SDC_FAULTS".Carrier_Fault[42] = 187;
END_REGION

REGION Network 71: CARRIER MOTION OFF FAULT
   RUNG wire#powerrail
      Contact( "EMS".Carrier[42].SDC_OUT.Faults.MotionOffFault )
      Coil( "DB302_HMI_Faults".Carrier42_Faults_2.%X0 )
   END_RUNG
   // the same network as SCL:
   "DB302_HMI_Faults".Carrier42_Faults_2.%X0 := "EMS".Carrier[42].SDC_OUT.Faults.MotionOffFault;
END_REGION

REGION Network 72: CARRIER MOTION ON FAULT
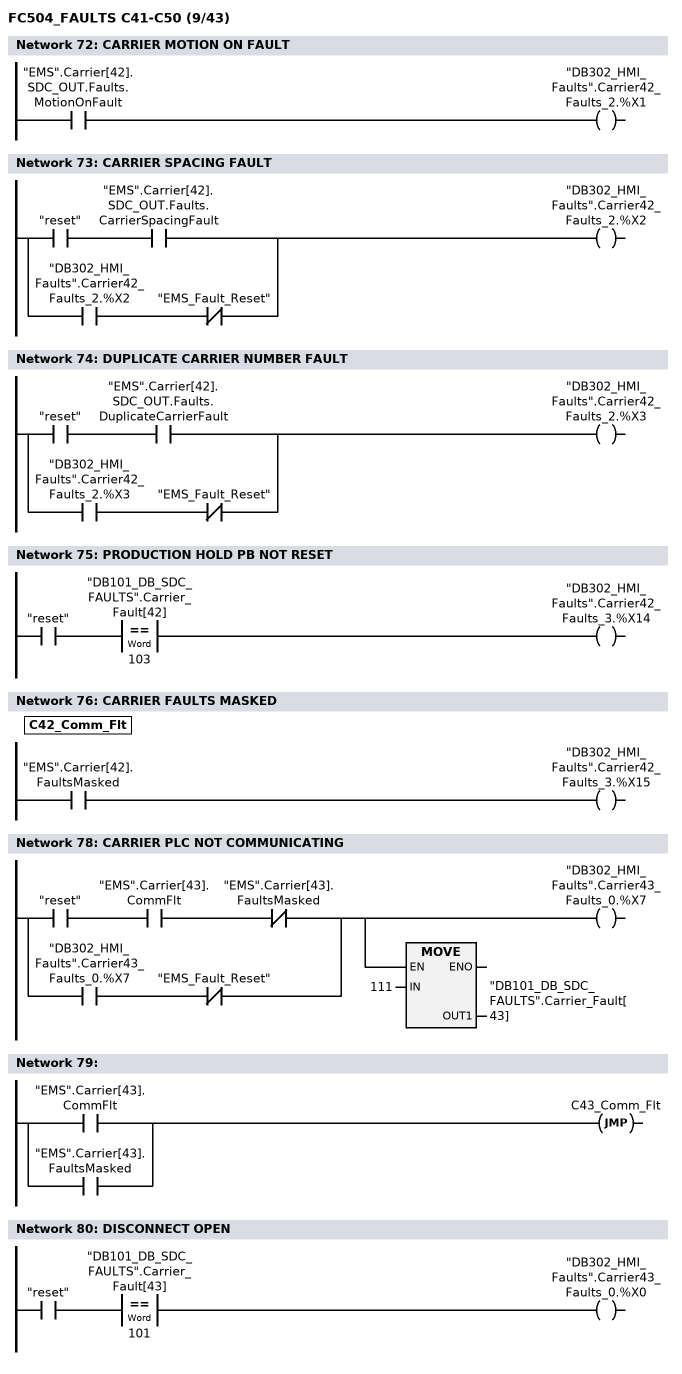
   RUNG wire#powerrail
      Contact( "EMS".Carrier[42].SDC_OUT.Faults.MotionOnFault )
      Coil( "DB302_HMI_Faults".Carrier42_Faults_2.%X1 )
   END_RUNG
   // the same network as SCL:
   "DB302_HMI_Faults".Carrier42_Faults_2.%X1 := "EMS".Carrier[42].SDC_OUT.Faults.MotionOnFault;
END_REGION

REGION Network 73: CARRIER SPACING FAULT
   RUNG wire#powerrail
      Contact( "reset" )
      Contact( "EMS".Carrier[42].SDC_OUT.Faults.CarrierSpacingFault )
      wire#w1
      Coil( "DB302_HMI_Faults".Carrier42_Faults_2.%X2 )
   END_RUNG
   RUNG wire#powerrail
      Contact( "DB302_HMI_Faults".Carrier42_Faults_2.%X2 )
      I_Contact( "EMS_Fault_Reset" )
   END_RUNG wire#w1
   // the same network as SCL:
   "DB302_HMI_Faults".Carrier42_Faults_2.%X2 := ("reset" AND "EMS".Carrier[42].SDC_OUT.Faults.CarrierSpacingFault) OR ("DB302_HMI_Faults".Carrier42_Faults_2.%X2 AND NOT "EMS_Fault_Reset");
END_REGION

REGION Network 74: DUPLICATE CARRIER NUMBER FAULT
   RUNG wire#powerrail
      Contact( "reset" )
      Contact( "EMS".Carrier[42].SDC_OUT.Faults.DuplicateCarrierFault )
      wire#w1
      Coil( "DB302_HMI_Faults".Carrier42_Faults_2.%X3 )
   END_RUNG
   RUNG wire#powerrail
      Contact( "DB302_HMI_Faults".Carrier42_Faults_2.%X3 )
      I_Contact( "EMS_Fault_Reset" )
   END_RUNG wire#w1
   // the same network as SCL:
   "DB302_HMI_Faults".Carrier42_Faults_2.%X3 := ("reset" AND "EMS".Carrier[42].SDC_OUT.Faults.DuplicateCarrierFault) OR ("DB302_HMI_Faults".Carrier42_Faults_2.%X3 AND NOT "EMS_Fault_Reset");
END_REGION

REGION Network 75: PRODUCTION HOLD PB NOT RESET
   RUNG wire#powerrail
      Contact( "reset" )
      { S7_Templates := "SrcType := Word" } EQ_Contact(in1 := "DB101_DB_SDC_FAULTS".Carrier_Fault[42], in2 := 103)
      Coil( "DB302_HMI_Faults".Carrier42_Faults_3.%X14 )
   END_RUNG
   // the same network as SCL:
   "DB302_HMI_Faults".Carrier42_Faults_3.%X14 := "reset" AND ("DB101_DB_SDC_FAULTS".Carrier_Fault[42] = 103);
END_REGION

REGION Network 76: CARRIER FAULTS MASKED
   Label( C42_Comm_Flt )
   RUNG wire#powerrail
      Contact( "EMS".Carrier[42].FaultsMasked )
      Coil( "DB302_HMI_Faults".Carrier42_Faults_3.%X15 )
   END_RUNG
   // the same network as SCL:
   C42_Comm_Flt:
   "DB302_HMI_Faults".Carrier42_Faults_3.%X15 := "EMS".Carrier[42].FaultsMasked;
END_REGION

REGION Network 77: CARRIER 43 FAULTS
END_REGION

REGION Network 78: CARRIER PLC NOT COMMUNICATING
   RUNG wire#powerrail
      Contact( "reset" )
      Contact( "EMS".Carrier[43].CommFlt )
      I_Contact( "EMS".Carrier[43].FaultsMasked )
      wire#w1
      Coil( "DB302_HMI_Faults".Carrier43_Faults_0.%X7 )
   END_RUNG
   RUNG wire#powerrail
      Contact( "DB302_HMI_Faults".Carrier43_Faults_0.%X7 )
      I_Contact( "EMS_Fault_Reset" )
   END_RUNG wire#w1
   RUNG wire#w1
      Move(in := 111, out1 => "DB101_DB_SDC_FAULTS".Carrier_Fault[43])
   END_RUNG
   // the same network as SCL:
   "DB302_HMI_Faults".Carrier43_Faults_0.%X7 := ("reset" AND "EMS".Carrier[43].CommFlt AND NOT "EMS".Carrier[43].FaultsMasked) OR ("DB302_HMI_Faults".Carrier43_Faults_0.%X7 AND NOT "EMS_Fault_Reset");
   IF "DB302_HMI_Faults".Carrier43_Faults_0.%X7 THEN "DB101_DB_SDC_FAULTS".Carrier_Fault[43] := 111; END_IF;
END_REGION

REGION Network 79
   RUNG wire#powerrail
      Contact( "EMS".Carrier[43].CommFlt )
      wire#w1
      JumpCoil( C43_Comm_Flt )
   END_RUNG
   RUNG wire#powerrail
      Contact( "EMS".Carrier[43].FaultsMasked )
   END_RUNG wire#w1
   // the same network as SCL:
   IF "EMS".Carrier[43].CommFlt OR "EMS".Carrier[43].FaultsMasked THEN GOTO C43_Comm_Flt; END_IF;
END_REGION

REGION Network 80: DISCONNECT OPEN
   RUNG wire#powerrail
      Contact( "reset" )
      { S7_Templates := "SrcType := Word" } EQ_Contact(in1 := "DB101_DB_SDC_FAULTS".Carrier_Fault[43], in2 := 101)
      Coil( "DB302_HMI_Faults".Carrier43_Faults_0.%X0 )
   END_RUNG
   // the same network as SCL:
   "DB302_HMI_Faults".Carrier43_Faults_0.%X0 := "reset" AND ("DB101_DB_SDC_FAULTS".Carrier_Fault[43] = 101);
END_REGION

REGION Network 81: PROFINET FAULT